// TIA Portal project "HEAT-1-CADIZ-V24" (V20)

(* hardware
DEVICE "S7-1200 station_1"  S7-1200 Station
   slot 0: "Rack_0"  S7-1200 Rack  Rack  V1.0
   slot 1: "PLC_1"  CPU 1214FC DC/DC/RLY  6ES7 214-1HF40-0XB0  V4.6
   slot 2: "DI 16x24VDC_1"  6ES7 221-1BH32-0XB0  V2.0
   slot 3: "DQ 16xRelay_1"  SM 1222 DQ16 x relay  6ES7 222-1HH32-0XB0  V2.0
   slot 4: "F-DI 8/16x24VDC_1"  SM 1226 F-DI8/16 x 24VDC  6ES7 226-6BA32-0XB0  V2.0
   slot 5: "F-DI 8/16x24VDC_2"  SM 1226 F-DI8/16 x 24VDC  6ES7 226-6BA32-0XB0  V2.0
   slot 6: "F-DQ 4x24VDC_1"  SM 1226 F-DQ4 x 24VDC  6ES7 226-6DA32-0XB0  V2.0
DEVICE "GSD device_1"  GSD.Device.PN
   slot 0: "Rack"  Rack  V1.0
   slot 0: "KRC5"  KUKA.PROFINET 6.0  0x300  V6.0
      slot 0: "KUKA.PROFINET 6.0"  KUKA.PROFINET 6.0
      slot 1: "Interface1"  Interface1
         slot 1: "Port001(XF3)"  Port001(XF3)
         slot 2: "Port002(XF4)"  Port002(XF4)
         slot 3: "Port003(XF5)"  Port003(XF5)
         slot 4: "Port004(XF6)"  Port004(XF6)
   slot 1: "64 safe digital in- and outputs (2.4)_1"  64 safe digital in- and outputs (2.4)  KUKADevF64_2.4
      slot 0: "64 safe digital in- and outputs (2.4)"  64 safe digital in- and outputs (2.4)
   slot 2: "1024 digital in- and outputs_1"  1024 digital in- and outputs  KUKA Device IO1024
      slot 0: "1024 digital in- and outputs"  1024 digital in- and outputs
DEVICE "HMI_1"  KTP1200 Basic PN
   slot 0: "HMI_1"  KTP1200 Basic PN  6AV2 123-2MB03-0AX0  17.0.0.0
   slot 1: "HMI_RT_1"  KTP1200 Basic PN  6AV2 123-2MB03-0AX0  17.0.0.0
   slot 5: "HMI_1.IE_CP_1"  PROFINET Interface  17.0.0.0
      slot 1: "PROFINET Interface_1"  PROFINET Interface
         slot 1: "Port_1"  Port
DEVICE "ET 200SP station_2"  ET 200SP-Station
   slot 0: "Rack_0"  Rack  6ES5 710-8MAx1
   slot 0: "islaparking"  IM 155-6 PN ST  6ES7 155-6AU01-0BN0  V4.2
   slot 1: "DI 16x24VDC ST_1"  DI 16x24VDC ST  6ES7 131-6BH01-0BA0  V0.0
      slot 1: "DI 16x24VDC ST_1"  DI 16x24VDC ST
   slot 2: "DI 8x24VDC ST_1"  DI 8x24VDC ST  6ES7 131-6BF01-0BA0  V0.0
      slot 1: "DI 8x24VDC ST_1"  DI 8x24VDC ST
   slot 3: "DQ 16x24VDC/0.5A ST_1"  DQ 16x24VDC/0.5A ST  6ES7 132-6BH01-0BA0  V0.0
      slot 1: "DQ 16x24VDC/0.5A ST_1"  DQ 16x24VDC/0.5A ST
   slot 4: "DQ 8x24VDC/0.5A ST_1"  DQ 8x24VDC/0.5A ST  6ES7 132-6BF01-0BA0  V0.0
      slot 1: "DQ 8x24VDC/0.5A ST_1"  DQ 8x24VDC/0.5A ST
   slot 5: "Server module_1"  Server module  6ES7 193-6PA00-0AA0  V1.1
      slot 1: "Server module_1"  Server module
   slot 127: "BA 2xRJ45"  BA 2xRJ45  6ES7 193-6AR00-0AA0  V0.0
      slot 1: "Port_1"  X1 P1R  6ES7 193-6AR00-0AA0  V0.0
      slot 2: "Port_2"  X1 P2R  6ES7 193-6AR00-0AA0  V0.0
DEVICE "ET 200SP station_1"  ET 200SP-Station
   slot 0: "Rack_0"  Rack  6ES5 710-8MAx1
   slot 0: "islarobot"  IM 155-6 PN ST  6ES7 155-6AU01-0BN0  V4.2
   slot 1: "DI 16x24VDC ST_1"  DI 16x24VDC ST  6ES7 131-6BH01-0BA0  V0.0
      slot 1: "DI 16x24VDC ST_1"  DI 16x24VDC ST
   slot 2: "DI 8x24VDC ST_1"  DI 8x24VDC ST  6ES7 131-6BF01-0BA0  V0.0
      slot 1: "DI 8x24VDC ST_1"  DI 8x24VDC ST
   slot 3: "DQ 16x24VDC/0.5A ST_1"  DQ 16x24VDC/0.5A ST  6ES7 132-6BH01-0BA0  V0.0
      slot 1: "DQ 16x24VDC/0.5A ST_1"  DQ 16x24VDC/0.5A ST
   slot 4: "DQ 8x24VDC/0.5A ST_1"  DQ 8x24VDC/0.5A ST  6ES7 132-6BF01-0BA0  V0.0
      slot 1: "DQ 8x24VDC/0.5A ST_1"  DQ 8x24VDC/0.5A ST
   slot 5: "Server module_1"  Server module  6ES7 193-6PA00-0AA0  V1.1
      slot 1: "Server module_1"  Server module
   slot 127: "BA 2xRJ45"  BA 2xRJ45  6ES7 193-6AR00-0AA0  V0.0
      slot 1: "Port_1"  X1 P1R  6ES7 193-6AR00-0AA0  V0.0
      slot 2: "Port_2"  X1 P2R  6ES7 193-6AR00-0AA0  V0.0
DEVICE "GSD device_2"  GSD.Device.PN
   slot 0: "Rack"  Rack  V1.0
   slot 0: "CPX"  CPX Rev 50  TN 197330
      slot 0: "CPX Rev 50"  CPX Rev 50
      slot 1: "PN-IO Interface"  PN-IO Interface
         slot 1: "Port 1"  Port 1
         slot 2: "Port 2"  Port 2
   slot 1: "FB43 PNIO Module_1"  FB43 PNIO Module  TN 8110369, CPX-FB43
      slot 0: "FB43 PNIO Module"  FB43 PNIO Module
   slot 2: "MPAL DIL 4 [32DO]_1"  MPAL DIL 4 [32DO]
      slot 0: "MPAL DIL 4 [32DO]"  MPAL DIL 4 [32DO]
DEVICE "ET 200SP station_3"  ET 200SP-Station
   slot 0: "Rack_0"  Rack  6ES5 710-8MAx1
   slot 0: "sistemadeagua"  IM 155-6 PN ST  6ES7 155-6AU01-0BN0  V4.2
   slot 1: "DI 8x24VDC ST_1"  DI 8x24VDC ST  6ES7 131-6BF01-0BA0  V0.0
      slot 1: "DI 8x24VDC ST_1"  DI 8x24VDC ST
   slot 2: "DQ 8x24VDC/0.5A ST_1"  DQ 8x24VDC/0.5A ST  6ES7 132-6BF01-0BA0  V0.0
      slot 1: "DQ 8x24VDC/0.5A ST_1"  DQ 8x24VDC/0.5A ST
   slot 3: "AI 4xU/I 2-wire ST_1"  AI 4xU/I 2-wire ST  6ES7 134-6HD01-0BA1  V2.0
      slot 1: "AI 4xU/I 2-wire ST_1"  AI 4xU/I 2-wire ST
   slot 4: "Server module_1"  Server module  6ES7 193-6PA00-0AA0  V1.1
      slot 1: "Server module_1"  Server module
   slot 127: "BA 2xRJ45"  BA 2xRJ45  6ES7 193-6AR00-0AA0  V0.0
      slot 1: "Port_1"  X1 P1R  6ES7 193-6AR00-0AA0  V0.0
      slot 2: "Port_2"  X1 P2R  6ES7 193-6AR00-0AA0  V0.0
DEVICE "GSD device_3"  GSD.Device.PN
   slot 0: "Rack"  Rack  V1.0
   slot 0: "CPX_1"  CPX Rev 50  TN 197330
      slot 0: "CPX Rev 50"  CPX Rev 50
      slot 1: "PN-IO Interface"  PN-IO Interface
         slot 1: "Port 1"  Port 1
         slot 2: "Port 2"  Port 2
   slot 1: "FB43 PNIO Module_1"  FB43 PNIO Module  TN 8110369, CPX-FB43
      slot 0: "FB43 PNIO Module"  FB43 PNIO Module
   slot 2: "16DI [16DI]_1"  16DI [16DI]
      slot 0: "16DI [16DI]"  16DI [16DI]
   slot 3: "16DI [16DI]_2"  16DI [16DI]
      slot 0: "16DI [16DI]"  16DI [16DI]
   slot 4: "MPAL DIL 4 [32DO]_1"  MPAL DIL 4 [32DO]
      slot 0: "MPAL DIL 4 [32DO]"  MPAL DIL 4 [32DO]
*)

// ===== PLC "PLC_1"  CPU 1214FC DC/DC/RLY =====

VAR_GLOBAL   // PLC tag table "Default tag table"
   "RES1 (reservado)" AT %Q500.0 : Bool;
   "eStopButtonCabinet" AT %I40.0 : Bool;   // Emergency-Stop cabinet — 1oo2 result
   "eStopButtonTank" AT %I40.1 : Bool;   // Emergency-Stop tank — 1oo2 result
   "eStopButtonTankPartnerCh" AT %I41.1 : Bool;   // partner channel 1oo2 — do not use
   "eStopButtonWaterSystem" AT %I40.2 : Bool;   // Emergency-Stop water system — 1oo2 result
   "eStopButtonWaterSystemPartnerCh" AT %I41.2 : Bool;   // partner channel 1oo2 — do not use
   "eStopButtonHmiPanel" AT %I40.3 : Bool;   // Emergency-Stop HMI panel — 1oo2 result
   "eStopButtonHmiPanelPartnerCh" AT %I41.3 : Bool;   // partner channel 1oo2 — do not use
   "eStopButtonLightCurtain1" AT %I40.4 : Bool;   // Emergency-Stop light curtain 1 — 1oo2 resul
   "eStopButtonLightCurtain1PartnerCh" AT %I41.4 : Bool;   // partner channel 1oo2 — do not use
   "eStopButtonDoor" AT %I40.5 : Bool;   // Emergency-Stop Door — 1oo2 result
   "eStopButtonDoorPartnerCh" AT %I41.5 : Bool;   // partner channel 1oo2 — do not use
   "lightCurtain1Ossd1" AT %I50.0 : Bool;   // Z2 – LC 1 OSSD 1 (receiver)
   "lightCurtain1Ossd2" AT %I51.0 : Bool;   // Z2 – LC 1 OSSD 2 (receiver)
   "lightCurtain3Ossd1" AT %I50.1 : Bool;   // Z2 – LC 3 OSSD 1 (receiver)
   "lightCurtain3Ossd2" AT %I51.1 : Bool;   // Z2 – LC 3 OSSD 2 (receiver)
   "lightCurtain6Ossd1" AT %I50.2 : Bool;   // Z2 – LC 6 OSSD 1 (receiver)
   "lightCurtain6Ossd2" AT %I51.2 : Bool;   // Z2 – LC 6 OSSD 2 (receiver)
   "enableAccessReqSelector" AT %I50.3 : Bool;   // Rotary selector – enabless request access
   "DoorClosedCh1" AT %I50.6 : Bool;   // Safety door closed interlock – contact 1
   "resetDoorButton" AT %I50.7 : Bool;   // Reset push‑button
   "SAF_DOOR_CLSD_CH2" AT %I51.6 : Bool;   // Safety door closed interlock – contact 2
   "SAF_DOOR_UNLOCK_CH1" AT %Q60.0 : Bool;   // Unlock safety door – redundant output 1
   "SAF_GATE_UNLOCK_CH2" AT %Q60.2 : Bool;   // Unlock safety door – redundant output 2
   "IND_RESET_LAMP" AT %Q10.0 : Bool;   // Reset indicator lamp
   "IND_STATUS_LAMP" AT %Q10.1 : Bool;   // System-status pilot light
   "CMD_PRESS_EXH_VALVE" AT %Q11.0 : Bool;   // Pressure/exhaust solenoid-valve command
   "STS_RECIRC_PUMP" AT %I20.0 : Bool;   // Recirculation-pump feedback
   "STS_TRANSFER_PUMP" AT %I20.1 : Bool;   // Transfer-pump feedback
   "ALM_UV_FILTER" AT %I20.2 : Bool;   // UV-filter fault alarm
   "ALM_PIT_LVL_LOW" AT %I20.3 : Bool;   // Sump low-level alarm
   "ALM_TANK_LVL_LOW" AT %I20.4 : Bool;   // Tank low-level alarm
   "STS_TANK_FILLING" AT %I20.5 : Bool;   // Tank filling status
   "STS_TANK_DRAINING" AT %I20.6 : Bool;   // Tank draining status
   "MODE_WATER_AUTO" AT %Q30.3 : Bool;   // CONMUTADOR AUTO
   "IND_BEACON2_GREEN" AT %Q30.4 : Bool;   // Beacon 2 – green
   "IND_BEACON2_RED" AT %Q30.5 : Bool;   // Beacon 2 – red
   "robotPresenceSignalZone1" AT %I500.0 : Bool;
   "robotPresenceSignalZone2" AT %I500.1 : Bool;
   "robotPresenceSignalZone3" AT %I500.2 : Bool;
   "eStopButtonCabinetPartnerCh" AT %I41.0 : Bool;   // partner channel 1oo2 — do not use
   "lightCurtain2Ossd1" AT %I300.0 : Bool;
   "lightCurtain2Ossd2" AT %I300.4 : Bool;
   "eStopButtonIslandRightPartner" AT %I300.5 : Bool;
   "lightCurtain4Ossd1" AT %I350.0 : Bool;
   "eStopButtonIslandLeft" AT %I350.1 : Bool;
   "lightCurtain5Ossd1" AT %I350.2 : Bool;
   "eStopButtonIslandLefttPartner" AT %I350.3 : Bool;   // partner channel 1oo2 — do not use
   "lightCurtain4Ossd2" AT %I350.4 : Bool;
   "lightCurtain5Ossd2" AT %I350.6 : Bool;
   "accessReqButtonZone2" AT %I51.4 : Bool;   // Illuminated push-button – access request for zone 2
   "accessReqButtonZone3" AT %I51.5 : Bool;   // Illuminated push-button – access request for zone 3
   "accessReqButtonZone1" AT %I51.3 : Bool;   // Illuminated push-button – access request for zone 1
   "eStopButtonIslandRight" AT %I300.1 : Bool;
   "NHE – E‑Stop externo  NO pulsado" AT %Q500.1 : Bool;
   "BS – Puerta cerrada" AT %Q500.2 : Bool;
   "QBS – Ack puerta" AT %Q500.3 : Bool;
   "SHS1 – Stop 1" AT %Q500.4 : Bool;
   "SHS2 – Stop 2" AT %Q500.5 : Bool;
   "RES6" AT %Q500.6 : Bool;
   "RES7" AT %Q500.7 : Bool;
   "US2 – 24 V US2" AT %Q501.0 : Bool;
   "SBH – Safe Op Stop" AT %Q501.1 : Bool;
   "RES11" AT %Q501.2 : Bool;
   "RES12" AT %Q501.3 : Bool;
   "RES13" AT %Q501.4 : Bool;
   "RES14" AT %Q501.5 : Bool;
   "RES15" AT %Q501.6 : Bool;
   "SPA – Power‑down Ack" AT %Q501.7 : Bool;
   "resetHmiButton" AT %I51.7 : Bool;
   "Tag_1" AT %M200.0 : Bool;
   "Tag_2" AT %M201.0 : Bool;
   "Tag_3" AT %M500.1 : Bool;
   "Tag_4" AT %M755.5 : Bool;
   "V5" AT %Q0.4 : Bool;   // Biestable_B_RETROCESO
   "ABRIR_TAPA_PEPA" AT %Q170.2 : Bool;
   "CERRAR_TAPA_PEPA" AT %Q170.3 : Bool;
   "ABRIR_TAPA_INMERSION" AT %Q170.4 : Bool;
   "CERRAR_TAPA_INMERSION" AT %Q170.5 : Bool;
   "ABRIR_TAPA_MARCADOR" AT %Q170.6 : Bool;
   "CERRAR_TAPA_MARCADOR" AT %Q170.7 : Bool;
   "ABRIR_TAPA_PERFILOMETRO" AT %Q171.0 : Bool;
   "CERRAR_TAPA_PERFILOMETRO" AT %Q171.1 : Bool;
   "V6" AT %Q0.5 : Bool;   // Biestable_A_AVANCE
   "V7" AT %Q0.6 : Bool;
   "V8" AT %Q0.7 : Bool;
   "moveCode_00" AT %Q616.0 : Bool;
   "goTrigger" AT %Q622.0 : Bool;
   "baseReqId_00" AT %Q620.0 : Bool;
   "baseReqId_01" AT %Q620.1 : Bool;
   "baseReqId_02" AT %Q620.2 : Bool;
   "baseReqId_03" AT %Q620.3 : Bool;
   "baseReqId_04" AT %Q620.4 : Bool;
   "baseReqId_05" AT %Q620.5 : Bool;
   "baseReqId_06" AT %Q620.6 : Bool;
   "baseReqId_07" AT %Q620.7 : Bool;
   "baseReqId_08" AT %Q621.0 : Bool;
   "baseReqId_09" AT %Q621.1 : Bool;
   "baseReqId_10" AT %Q621.2 : Bool;
   "baseReqId_11" AT %Q621.3 : Bool;
   "baseReqId_12" AT %Q621.4 : Bool;
   "baseReqId_13" AT %Q621.5 : Bool;
   "baseReqId_14" AT %Q621.6 : Bool;
   "baseReqId_15" AT %Q621.7 : Bool;
   "moveCode_01" AT %Q616.1 : Bool;
   "moveCode_02" AT %Q616.2 : Bool;
   "moveCode_03" AT %Q616.3 : Bool;
   "moveCode_04" AT %Q616.4 : Bool;
   "moveCode_05" AT %Q616.5 : Bool;
   "moveCode_06" AT %Q616.6 : Bool;
   "moveCode_07" AT %Q616.7 : Bool;
   "moveCode_08" AT %Q617.0 : Bool;
   "moveCode_09" AT %Q617.1 : Bool;
   "moveCode_10" AT %Q617.2 : Bool;
   "moveCode_11" AT %Q617.3 : Bool;
   "moveCode_12" AT %Q617.4 : Bool;
   "moveCode_13" AT %Q617.5 : Bool;
   "moveCode_14" AT %Q617.6 : Bool;
   "moveCode_15" AT %Q617.7 : Bool;
   "toolNo_00" AT %I625.0 : Bool;
   "toolNo_01" AT %I625.1 : Bool;
   "toolNo_02" AT %I625.2 : Bool;
   "toolNo_03" AT %I625.3 : Bool;
   "toolNo_04" AT %I625.4 : Bool;
   "toolNo_05" AT %I625.5 : Bool;
   "toolNo_06" AT %I625.6 : Bool;
   "toolNo_07" AT %I625.7 : Bool;
   "baseNo_00" AT %I626.0 : Bool;
   "baseNo_01" AT %I626.1 : Bool;
   "baseNo_02" AT %I626.2 : Bool;
   "baseNo_03" AT %I626.3 : Bool;
   "baseNo_04" AT %I626.4 : Bool;
   "baseNo_05" AT %I626.5 : Bool;
   "baseNo_06" AT %I626.6 : Bool;
   "baseNo_07" AT %I626.7 : Bool;
   "toolNoByte" AT %IB625 : Byte;
   "baseNoByte" AT %IB626 : Byte;
   "programReqId_00" AT %Q623.0 : Bool;
   "programReqId_01" AT %Q623.1 : Bool;
   "programReqId_02" AT %Q623.2 : Bool;
   "programReqId_03" AT %Q623.3 : Bool;
   "programReqId_04" AT %Q623.4 : Bool;
   "programReqId_05" AT %Q623.5 : Bool;
   "programReqId_06" AT %Q623.6 : Bool;
   "programReqId_07" AT %Q623.7 : Bool;
   "programReqId_08" AT %Q624.0 : Bool;
   "programReqId_09" AT %Q624.1 : Bool;
   "programReqId_10" AT %Q624.2 : Bool;
   "programReqId_11" AT %Q624.3 : Bool;
   "programReqId_12" AT %Q624.4 : Bool;
   "programReqId_13" AT %Q624.5 : Bool;
   "programReqId_14" AT %Q624.6 : Bool;
   "programReqId_15" AT %Q624.7 : Bool;
   "programReqId" AT %QW623 : Word;
   "PRUEBA_4" AT %Q4.4 : Bool;
   "PRUEBA_5" AT %Q4.5 : Bool;
   "PRUEBA_JOAQUIN" AT %Q4.0 : Bool;
   "PRUEBA_6" AT %Q4.6 : Bool;
   "PRUEBA_7" AT %Q4.7 : Bool;
   "cancelGo" AT %Q625.0 : Bool;
   "pauseGo" AT %Q625.1 : Bool;
   "resumeGo" AT %Q625.2 : Bool;
   "ACTIVAR_AGUA" AT %Q220.1 : Bool;   // VALVULA EMBARCADA ISLA ROBOT
   "AGUA_JOAQUIN" AT %Q4.3 : Bool;   // SISTEMA DE AGUA - JOAQUIN
   "PGNO_BIT_00" AT %Q626.0 : Bool;   // $IN[209] en KUKA
   "PGNO_BIT_01" AT %Q626.1 : Bool;   // $IN[210] en KUKA
   "PGNO_BIT_02" AT %Q626.2 : Bool;   // $IN[211] en KUKA
   "PGNO_BIT_03" AT %Q626.3 : Bool;
   "PGNO_BIT_04" AT %Q626.4 : Bool;
   "PGNO_BIT_05" AT %Q626.5 : Bool;
   "PGNO_BIT_06" AT %Q626.6 : Bool;
   "PGNO_BIT_07" AT %Q626.7 : Bool;
   "PGNO_PARITY" AT %Q627.0 : Bool;   // $IN[217] en KUKA
   "PGNO_VALID" AT %Q627.1 : Bool;   // $IN[218] en KUKA
   "$EXT_START" AT %Q627.2 : Bool;   // $IN[219] en KUKA
   "$MOVE_ENABLE" AT %Q627.3 : Bool;   // $IN[220] en KUKA
   "$CONF_MESS" AT %Q627.4 : Bool;   // $IN[221] en KUKA
   "$DRIVES_OFF" AT %Q627.5 : Bool;   // $IN[222] en KUKA
   "$DRIVES_ON" AT %Q627.6 : Bool;   // $IN[223] en KUKA
   "$I_O_ACT" AT %Q627.7 : Bool;   // $IN[224] en KUKA
   "PGNO_REQ" AT %I624.7 : Bool;   // OUT[200] EN KUKA
   "startAutoExt" AT %M777.0 : Bool;
   "Tag_6" AT %Q220.0 : Bool;
   "Tag_7" AT %Q4.1 : Bool;
   "Tag_8" AT %Q4.2 : Bool;
   "Tag_9" AT %I0.4 : Bool;
   "Tag_10" AT %I0.0 : Bool;
   "Tag_11" AT %I0.1 : Bool;
   "Tag_12" AT %I0.2 : Bool;
   "Tag_13" AT %I0.3 : Bool;
   "Tag_14" AT %I210.1 : Bool;
   "Tag_15" AT %I210.2 : Bool;
   "Tag_16" AT %I210.0 : Bool;
   "Tag_17" AT %I210.3 : Bool;
   "Tag_18" AT %I210.4 : Bool;
   "AchimHmiEnable" AT %M202.0 : Bool;
   "toolIdProxy1" AT %I201.3 : Bool;
   "toolIdProxy2" AT %I201.2 : Bool;
   "toolIdProxy3" AT %I201.1 : Bool;
   "toolIdProxy4" AT %I201.0 : Bool;
   "dockValveV2UnlockOnPole" AT %Q171.6 : Bool;
   "$PRO_ACT" AT %I627.2 : Bool;   // OUT[219] EN KUKA
   "$STOPMESS" AT %I627.1 : Bool;   // OUT[218] EN KUKA
   "$PERI_RDY" AT %I627.0 : Bool;   // OUT[217] EN KUKA
   "robotInLoopKukaControl" AT %Q628.0 : Bool;
   "robotInLoopSupervisor" AT %Q628.1 : Bool;
   "xInicial_00" AT %Q632.0 : Bool;
   "xInicial_01" AT %Q632.1 : Bool;
   "xInicial_02" AT %Q632.2 : Bool;
   "xInicial_03" AT %Q632.3 : Bool;
   "xInicial_04" AT %Q632.4 : Bool;
   "xInicial_05" AT %Q632.5 : Bool;
   "xInicial_06" AT %Q632.6 : Bool;
   "xInicial_07" AT %Q632.7 : Bool;
   "xInicial_08" AT %Q633.0 : Bool;
   "xInicial_09" AT %Q633.1 : Bool;
   "xInicial_10" AT %Q633.2 : Bool;
   "xInicial_11" AT %Q633.3 : Bool;
   "xInicial_12" AT %Q633.4 : Bool;
   "xInicial_13" AT %Q633.5 : Bool;
   "xInicial_14" AT %Q633.6 : Bool;
   "xInicial_15" AT %Q633.7 : Bool;
   "xInicial_16" AT %Q634.0 : Bool;
   "xInicial_17" AT %Q634.1 : Bool;
   "xInicial_18" AT %Q634.2 : Bool;
   "xInicial_19" AT %Q634.3 : Bool;
   "xInicial_20" AT %Q634.4 : Bool;
   "xInicial_21" AT %Q634.5 : Bool;
   "xInicial_22" AT %Q634.6 : Bool;
   "xInicial_23" AT %Q634.7 : Bool;
   "xInicial_24" AT %Q635.0 : Bool;
   "xInicial_25" AT %Q635.1 : Bool;
   "xInicial_26" AT %Q635.2 : Bool;
   "xInicial_27" AT %Q635.3 : Bool;
   "xInicial_28" AT %Q635.4 : Bool;
   "xInicial_29" AT %Q635.5 : Bool;
   "xInicial_30" AT %Q635.6 : Bool;
   "xInicial_31" AT %Q635.7 : Bool;
   "yInicial_00" AT %Q636.0 : Bool;
   "yInicial_01" AT %Q636.1 : Bool;
   "yInicial_02" AT %Q636.2 : Bool;
   "yInicial_03" AT %Q636.3 : Bool;
   "yInicial_04" AT %Q636.4 : Bool;
   "yInicial_05" AT %Q636.5 : Bool;
   "yInicial_06" AT %Q636.6 : Bool;
   "yInicial_07" AT %Q636.7 : Bool;
   "yInicial_08" AT %Q637.0 : Bool;
   "yInicial_09" AT %Q637.1 : Bool;
   "yInicial_10" AT %Q637.2 : Bool;
   "yInicial_11" AT %Q637.3 : Bool;
   "yInicial_12" AT %Q637.4 : Bool;
   "yInicial_13" AT %Q637.5 : Bool;
   "yInicial_14" AT %Q637.6 : Bool;
   "yInicial_15" AT %Q637.7 : Bool;
   "yInicial_16" AT %Q638.0 : Bool;
   "yInicial_17" AT %Q638.1 : Bool;
   "yInicial_18" AT %Q638.2 : Bool;
   "yInicial_19" AT %Q638.3 : Bool;
   "yInicial_20" AT %Q638.4 : Bool;
   "yInicial_21" AT %Q638.5 : Bool;
   "yInicial_22" AT %Q638.6 : Bool;
   "yInicial_23" AT %Q638.7 : Bool;
   "yInicial_24" AT %Q639.0 : Bool;
   "yInicial_25" AT %Q639.1 : Bool;
   "yInicial_26" AT %Q639.2 : Bool;
   "yInicial_27" AT %Q639.3 : Bool;
   "yInicial_28" AT %Q639.4 : Bool;
   "yInicial_29" AT %Q639.5 : Bool;
   "yInicial_30" AT %Q639.6 : Bool;
   "yInicial_31" AT %Q639.7 : Bool;
   "zInicial_00" AT %Q640.0 : Bool;
   "zInicial_01" AT %Q640.1 : Bool;
   "zInicial_02" AT %Q640.2 : Bool;
   "zInicial_03" AT %Q640.3 : Bool;
   "zInicial_04" AT %Q640.4 : Bool;
   "zInicial_05" AT %Q640.5 : Bool;
   "zInicial_06" AT %Q640.6 : Bool;
   "zInicial_07" AT %Q640.7 : Bool;
   "zInicial_08" AT %Q641.0 : Bool;
   "zInicial_09" AT %Q641.1 : Bool;
   "zInicial_10" AT %Q641.2 : Bool;
   "zInicial_11" AT %Q641.3 : Bool;
   "zInicial_12" AT %Q641.4 : Bool;
   "zInicial_13" AT %Q641.5 : Bool;
   "zInicial_14" AT %Q641.6 : Bool;
   "zInicial_15" AT %Q641.7 : Bool;
   "zInicial_16" AT %Q642.0 : Bool;
   "zInicial_17" AT %Q642.1 : Bool;
   "zInicial_18" AT %Q642.2 : Bool;
   "zInicial_19" AT %Q642.3 : Bool;
   "zInicial_20" AT %Q642.4 : Bool;
   "zInicial_21" AT %Q642.5 : Bool;
   "zInicial_22" AT %Q642.6 : Bool;
   "zInicial_23" AT %Q642.7 : Bool;
   "zInicial_24" AT %Q643.0 : Bool;
   "zInicial_25" AT %Q643.1 : Bool;
   "zInicial_26" AT %Q643.2 : Bool;
   "zInicial_27" AT %Q643.3 : Bool;
   "zInicial_28" AT %Q643.4 : Bool;
   "zInicial_29" AT %Q643.5 : Bool;
   "zInicial_30" AT %Q643.6 : Bool;
   "zInicial_31" AT %Q643.7 : Bool;
   "e1Inicial_00" AT %Q644.0 : Bool;
   "e1Inicial_01" AT %Q644.1 : Bool;
   "e1Inicial_02" AT %Q644.2 : Bool;
   "e1Inicial_03" AT %Q644.3 : Bool;
   "e1Inicial_04" AT %Q644.4 : Bool;
   "e1Inicial_05" AT %Q644.5 : Bool;
   "e1Inicial_06" AT %Q644.6 : Bool;
   "e1Inicial_07" AT %Q644.7 : Bool;
   "e1Inicial_08" AT %Q645.0 : Bool;
   "e1Inicial_09" AT %Q645.1 : Bool;
   "e1Inicial_10" AT %Q645.2 : Bool;
   "e1Inicial_11" AT %Q645.3 : Bool;
   "e1Inicial_12" AT %Q645.4 : Bool;
   "e1Inicial_13" AT %Q645.5 : Bool;
   "e1Inicial_14" AT %Q645.6 : Bool;
   "e1Inicial_15" AT %Q645.7 : Bool;
   "e1Inicial_16" AT %Q646.0 : Bool;
   "e1Inicial_17" AT %Q646.1 : Bool;
   "e1Inicial_18" AT %Q646.2 : Bool;
   "e1Inicial_19" AT %Q646.3 : Bool;
   "e1Inicial_20" AT %Q646.4 : Bool;
   "e1Inicial_21" AT %Q646.5 : Bool;
   "e1Inicial_22" AT %Q646.6 : Bool;
   "e1Inicial_23" AT %Q646.7 : Bool;
   "e1Inicial_24" AT %Q647.0 : Bool;
   "e1Inicial_25" AT %Q647.1 : Bool;
   "e1Inicial_26" AT %Q647.2 : Bool;
   "e1Inicial_27" AT %Q647.3 : Bool;
   "e1Inicial_28" AT %Q647.4 : Bool;
   "e1Inicial_29" AT %Q647.5 : Bool;
   "e1Inicial_30" AT %Q647.6 : Bool;
   "e1Inicial_31" AT %Q647.7 : Bool;
   "xFinal_00" AT %Q648.0 : Bool;
   "xFinal_01" AT %Q648.1 : Bool;
   "xFinal_02" AT %Q648.2 : Bool;
   "xFinal_03" AT %Q648.3 : Bool;
   "xFinal_04" AT %Q648.4 : Bool;
   "xFinal_05" AT %Q648.5 : Bool;
   "xFinal_06" AT %Q648.6 : Bool;
   "xFinal_07" AT %Q648.7 : Bool;
   "xFinal_08" AT %Q649.0 : Bool;
   "xFinal_09" AT %Q649.1 : Bool;
   "xFinal_10" AT %Q649.2 : Bool;
   "xFinal_11" AT %Q649.3 : Bool;
   "xFinal_12" AT %Q649.4 : Bool;
   "xFinal_13" AT %Q649.5 : Bool;
   "xFinal_14" AT %Q649.6 : Bool;
   "xFinal_15" AT %Q649.7 : Bool;
   "xFinal_16" AT %Q650.0 : Bool;
   "xFinal_17" AT %Q650.1 : Bool;
   "xFinal_18" AT %Q650.2 : Bool;
   "xFinal_19" AT %Q650.3 : Bool;
   "xFinal_20" AT %Q650.4 : Bool;
   "xFinal_21" AT %Q650.5 : Bool;
   "xFinal_22" AT %Q650.6 : Bool;
   "xFinal_23" AT %Q650.7 : Bool;
   "xFinal_24" AT %Q651.0 : Bool;
   "xFinal_25" AT %Q651.1 : Bool;
   "xFinal_26" AT %Q651.2 : Bool;
   "xFinal_27" AT %Q651.3 : Bool;
   "xFinal_28" AT %Q651.4 : Bool;
   "xFinal_29" AT %Q651.5 : Bool;
   "xFinal_30" AT %Q651.6 : Bool;
   "xFinal_31" AT %Q651.7 : Bool;
   "yFinal_00" AT %Q652.0 : Bool;
   "yFinal_01" AT %Q652.1 : Bool;
   "yFinal_02" AT %Q652.2 : Bool;
   "yFinal_03" AT %Q652.3 : Bool;
   "yFinal_04" AT %Q652.4 : Bool;
   "yFinal_05" AT %Q652.5 : Bool;
   "yFinal_06" AT %Q652.6 : Bool;
   "yFinal_07" AT %Q652.7 : Bool;
   "yFinal_08" AT %Q653.0 : Bool;
   "yFinal_09" AT %Q653.1 : Bool;
   "yFinal_10" AT %Q653.2 : Bool;
   "yFinal_11" AT %Q653.3 : Bool;
   "yFinal_12" AT %Q653.4 : Bool;
   "yFinal_13" AT %Q653.5 : Bool;
   "yFinal_14" AT %Q653.6 : Bool;
   "yFinal_15" AT %Q653.7 : Bool;
   "yFinal_16" AT %Q654.0 : Bool;
   "yFinal_17" AT %Q654.1 : Bool;
   "yFinal_18" AT %Q654.2 : Bool;
   "yFinal_19" AT %Q654.3 : Bool;
   "yFinal_20" AT %Q654.4 : Bool;
   "yFinal_21" AT %Q654.5 : Bool;
   "yFinal_22" AT %Q654.6 : Bool;
   "yFinal_23" AT %Q654.7 : Bool;
   "yFinal_24" AT %Q655.0 : Bool;
   "yFinal_25" AT %Q655.1 : Bool;
   "yFinal_26" AT %Q655.2 : Bool;
   "yFinal_27" AT %Q655.3 : Bool;
   "yFinal_28" AT %Q655.4 : Bool;
   "yFinal_29" AT %Q655.5 : Bool;
   "yFinal_30" AT %Q655.6 : Bool;
   "yFinal_31" AT %Q655.7 : Bool;
   "zFinal_00" AT %Q656.0 : Bool;
   "zFinal_01" AT %Q656.1 : Bool;
   "zFinal_02" AT %Q656.2 : Bool;
   "zFinal_03" AT %Q656.3 : Bool;
   "zFinal_04" AT %Q656.4 : Bool;
   "zFinal_05" AT %Q656.5 : Bool;
   "zFinal_06" AT %Q656.6 : Bool;
   "zFinal_07" AT %Q656.7 : Bool;
   "zFinal_08" AT %Q657.0 : Bool;
   "zFinal_09" AT %Q657.1 : Bool;
   "zFinal_10" AT %Q657.2 : Bool;
   "zFinal_11" AT %Q657.3 : Bool;
   "zFinal_12" AT %Q657.4 : Bool;
   "zFinal_13" AT %Q657.5 : Bool;
   "zFinal_14" AT %Q657.6 : Bool;
   "zFinal_15" AT %Q657.7 : Bool;
   "zFinal_16" AT %Q658.0 : Bool;
   "zFinal_17" AT %Q658.1 : Bool;
   "zFinal_18" AT %Q658.2 : Bool;
   "zFinal_19" AT %Q658.3 : Bool;
   "zFinal_20" AT %Q658.4 : Bool;
   "zFinal_21" AT %Q658.5 : Bool;
   "zFinal_22" AT %Q658.6 : Bool;
   "zFinal_23" AT %Q658.7 : Bool;
   "zFinal_24" AT %Q659.0 : Bool;
   "zFinal_25" AT %Q659.1 : Bool;
   "zFinal_26" AT %Q659.2 : Bool;
   "zFinal_27" AT %Q659.3 : Bool;
   "zFinal_28" AT %Q659.4 : Bool;
   "zFinal_29" AT %Q659.5 : Bool;
   "zFinal_30" AT %Q659.6 : Bool;
   "zFinal_31" AT %Q659.7 : Bool;
   "e1Final_00" AT %Q660.0 : Bool;
   "e1Final_01" AT %Q660.1 : Bool;
   "e1Final_02" AT %Q660.2 : Bool;
   "e1Final_03" AT %Q660.3 : Bool;
   "e1Final_04" AT %Q660.4 : Bool;
   "e1Final_05" AT %Q660.5 : Bool;
   "e1Final_06" AT %Q660.6 : Bool;
   "e1Final_07" AT %Q660.7 : Bool;
   "e1Final_08" AT %Q661.0 : Bool;
   "e1Final_09" AT %Q661.1 : Bool;
   "e1Final_10" AT %Q661.2 : Bool;
   "e1Final_11" AT %Q661.3 : Bool;
   "e1Final_12" AT %Q661.4 : Bool;
   "e1Final_13" AT %Q661.5 : Bool;
   "e1Final_14" AT %Q661.6 : Bool;
   "e1Final_15" AT %Q661.7 : Bool;
   "e1Final_16" AT %Q662.0 : Bool;
   "e1Final_17" AT %Q662.1 : Bool;
   "e1Final_18" AT %Q662.2 : Bool;
   "e1Final_19" AT %Q662.3 : Bool;
   "e1Final_20" AT %Q662.4 : Bool;
   "e1Final_21" AT %Q662.5 : Bool;
   "e1Final_22" AT %Q662.6 : Bool;
   "e1Final_23" AT %Q662.7 : Bool;
   "e1Final_24" AT %Q663.0 : Bool;
   "e1Final_25" AT %Q663.1 : Bool;
   "e1Final_26" AT %Q663.2 : Bool;
   "e1Final_27" AT %Q663.3 : Bool;
   "e1Final_28" AT %Q663.4 : Bool;
   "e1Final_29" AT %Q663.5 : Bool;
   "e1Final_30" AT %Q663.6 : Bool;
   "e1Final_31" AT %Q663.7 : Bool;
   "velRequest_00" AT %Q664.0 : Bool;
   "velRequest_01" AT %Q664.1 : Bool;
   "velRequest_02" AT %Q664.2 : Bool;
   "velRequest_03" AT %Q664.3 : Bool;
   "velRequest_04" AT %Q664.4 : Bool;
   "velRequest_05" AT %Q664.5 : Bool;
   "velRequest_06" AT %Q664.6 : Bool;
   "velRequest_07" AT %Q664.7 : Bool;
   "velRequest_08" AT %Q665.0 : Bool;
   "velRequest_09" AT %Q665.1 : Bool;
   "velRequest_10" AT %Q665.2 : Bool;
   "velRequest_11" AT %Q665.3 : Bool;
   "velRequest_12" AT %Q665.4 : Bool;
   "velRequest_13" AT %Q665.5 : Bool;
   "velRequest_14" AT %Q665.6 : Bool;
   "velRequest_15" AT %Q665.7 : Bool;
   "indexRequest_00" AT %Q666.0 : Bool;
   "indexRequest_01" AT %Q666.1 : Bool;
   "indexRequest_02" AT %Q666.2 : Bool;
   "indexRequest_03" AT %Q666.3 : Bool;
   "indexRequest_04" AT %Q666.4 : Bool;
   "indexRequest_05" AT %Q666.5 : Bool;
   "indexRequest_06" AT %Q666.6 : Bool;
   "indexRequest_07" AT %Q666.7 : Bool;
   "indexRequest_08" AT %Q667.0 : Bool;
   "indexRequest_09" AT %Q667.1 : Bool;
   "indexRequest_10" AT %Q667.2 : Bool;
   "indexRequest_11" AT %Q667.3 : Bool;
   "indexRequest_12" AT %Q667.4 : Bool;
   "indexRequest_13" AT %Q667.5 : Bool;
   "indexRequest_14" AT %Q667.6 : Bool;
   "indexRequest_15" AT %Q667.7 : Bool;
   "Tag_5" AT %M1000.1 : Bool;
   "toolInRobot_00" AT %Q668.0 : Bool;
   "toolInRobot_01" AT %Q668.1 : Bool;
   "toolInRobot_02" AT %Q668.2 : Bool;
   "toolInRobot_03" AT %Q668.3 : Bool;
   "toolInRobot_04" AT %Q668.4 : Bool;
   "toolInRobot_05" AT %Q668.5 : Bool;
   "toolInRobot_06" AT %Q668.6 : Bool;
   "toolInRobot_07" AT %Q668.7 : Bool;
   "kukaFeedBackToolInRobot" AT %QW668 : Word;
   "toolInRobot_08" AT %Q669.0 : Bool;
   "toolInRobot_09" AT %Q669.1 : Bool;
   "toolInRobot_10" AT %Q669.2 : Bool;
   "toolInRobot_11" AT %Q669.3 : Bool;
   "toolInRobot_12" AT %Q669.4 : Bool;
   "toolInRobot_13" AT %Q669.5 : Bool;
   "toolInRobot_14" AT %Q669.6 : Bool;
   "toolInRobot_15" AT %Q669.7 : Bool;
   "kukaAtPerspexPos" AT %I698.0 : Bool;
   "kukaAtGainPos" AT %I698.1 : Bool;
   "kukaAtTcgPos" AT %I698.2 : Bool;
   "kukaAtRefStart" AT %I698.3 : Bool;
   "kukaAtInspStart" AT %I698.4 : Bool;
   "kukaRefScanFin" AT %I698.5 : Bool;
   "kukaInspScanFin" AT %I698.6 : Bool;
   "requestVelocityKuka" AT %QW664 : Word;
   "requestIndexKuka" AT %QW666 : Word;
   "$IN_HOME" AT %I627.3 : Bool;   // OUT[220] EN KUKA
   "$EXT" AT %I627.4 : Bool;   // OUT[221] EN KUKA
END_VAR

VAR_GLOBAL   // PLC tag table "Robot Jog"
   "tcpTargetX_01" AT %Q600.1 : Bool;
   "tcpTargetX_02" AT %Q600.2 : Bool;
   "tcpTargetX_03" AT %Q600.3 : Bool;
   "tcpTargetX_04" AT %Q600.4 : Bool;
   "tcpTargetX_05" AT %Q600.5 : Bool;
   "tcpTargetX_08" AT %Q601.0 : Bool;
   "tcpTargetX_16" AT %Q602.0 : Bool;
   "tcpTargetX_17" AT %Q602.1 : Bool;
   "tcpTargetX_06" AT %Q600.6 : Bool;
   "tcpTargetX_07" AT %Q600.7 : Bool;
   "tcpTargetX_09" AT %Q601.1 : Bool;
   "tcpTargetX_10" AT %Q601.2 : Bool;
   "tcpTargetX_11" AT %Q601.3 : Bool;
   "tcpTargetX_12" AT %Q601.4 : Bool;
   "tcpTargetX_13" AT %Q601.5 : Bool;
   "tcpTargetX_14" AT %Q601.6 : Bool;
   "tcpTargetX_15" AT %Q601.7 : Bool;
   "tcpTargetX_18" AT %Q602.2 : Bool;
   "tcpTargetX_19" AT %Q602.3 : Bool;
   "tcpTargetX_20" AT %Q602.4 : Bool;
   "tcpTargetX_21" AT %Q602.5 : Bool;
   "tcpTargetX_22" AT %Q602.6 : Bool;
   "tcpTargetX_23" AT %Q602.7 : Bool;
   "tcpTargetX_24" AT %Q603.0 : Bool;
   "tcpTargetX_25" AT %Q603.1 : Bool;
   "tcpTargetX_26" AT %Q603.2 : Bool;
   "tcpTargetX_27" AT %Q603.3 : Bool;
   "tcpTargetX_28" AT %Q603.4 : Bool;
   "tcpTargetX_29" AT %Q603.5 : Bool;
   "tcpTargetX_30" AT %Q603.6 : Bool;
   "tcpTargetX_31" AT %Q603.7 : Bool;
   "tcpTargetY_00" AT %Q604.0 : Bool;
   "tcpTargetY_01" AT %Q604.1 : Bool;
   "tcpTargetY_02" AT %Q604.2 : Bool;
   "tcpTargetY_03" AT %Q604.3 : Bool;
   "tcpTargetY_04" AT %Q604.4 : Bool;
   "tcpTargetY_05" AT %Q604.5 : Bool;
   "tcpTargetY_06" AT %Q604.6 : Bool;
   "tcpTargetY_07" AT %Q604.7 : Bool;
   "tcpTargetY_08" AT %Q605.0 : Bool;
   "tcpTargetY_09" AT %Q605.1 : Bool;
   "tcpTargetY_10" AT %Q605.2 : Bool;
   "tcpTargetY_11" AT %Q605.3 : Bool;
   "tcpTargetY_12" AT %Q605.4 : Bool;
   "tcpTargetY_13" AT %Q605.5 : Bool;
   "tcpTargetY_14" AT %Q605.6 : Bool;
   "tcpTargetY_15" AT %Q605.7 : Bool;
   "tcpTargetY_16" AT %Q606.0 : Bool;   // $IN[49]
   "tcpTargetY_17" AT %Q606.1 : Bool;   // $IN[50]
   "tcpTargetY_18" AT %Q606.2 : Bool;   // $IN[51]
   "tcpTargetY_19" AT %Q606.3 : Bool;   // true
   "tcpTargetY_20" AT %Q606.4 : Bool;
   "tcpTargetY_21" AT %Q606.5 : Bool;   // true
   "tcpTargetY_22" AT %Q606.6 : Bool;   // true
   "tcpTargetY_23" AT %Q606.7 : Bool;   // true
   "tcpTargetY_24" AT %Q607.0 : Bool;   // true
   "tcpTargetY_25" AT %Q607.1 : Bool;   // true
   "tcpTargetY_26" AT %Q607.2 : Bool;   // true
   "tcpTargetY_27" AT %Q607.3 : Bool;
   "tcpTargetY_28" AT %Q607.4 : Bool;
   "tcpTargetY_29" AT %Q607.5 : Bool;
   "tcpTargetY_30" AT %Q607.6 : Bool;
   "tcpTargetY_31" AT %Q607.7 : Bool;
   "tcpTargetZ_00" AT %Q608.0 : Bool;
   "tcpTargetZ_01" AT %Q608.1 : Bool;
   "tcpTargetZ_02" AT %Q608.2 : Bool;
   "tcpTargetZ_03" AT %Q608.3 : Bool;
   "tcpTargetZ_04" AT %Q608.4 : Bool;
   "tcpTargetZ_05" AT %Q608.5 : Bool;
   "tcpTargetZ_06" AT %Q608.6 : Bool;
   "tcpTargetZ_07" AT %Q608.7 : Bool;
   "tcpTargetZ_08" AT %Q609.0 : Bool;
   "tcpTargetZ_09" AT %Q609.1 : Bool;
   "tcpTargetZ_10" AT %Q609.2 : Bool;
   "tcpTargetZ_11" AT %Q609.3 : Bool;
   "tcpTargetZ_12" AT %Q609.4 : Bool;
   "tcpTargetZ_13" AT %Q609.5 : Bool;
   "tcpTargetZ_14" AT %Q609.6 : Bool;
   "tcpTargetZ_15" AT %Q609.7 : Bool;
   "tcpTargetZ_16" AT %Q610.0 : Bool;
   "tcpTargetZ_17" AT %Q610.1 : Bool;
   "tcpTargetZ_18" AT %Q610.2 : Bool;
   "tcpTargetZ_19" AT %Q610.3 : Bool;
   "tcpTargetZ_20" AT %Q610.4 : Bool;
   "tcpTargetZ_21" AT %Q610.5 : Bool;
   "tcpTargetZ_22" AT %Q610.6 : Bool;
   "tcpTargetZ_23" AT %Q610.7 : Bool;
   "tcpTargetZ_24" AT %Q611.0 : Bool;
   "tcpTargetZ_25" AT %Q611.1 : Bool;
   "tcpTargetZ_26" AT %Q611.2 : Bool;
   "tcpTargetZ_27" AT %Q611.3 : Bool;
   "tcpTargetZ_28" AT %Q611.4 : Bool;
   "tcpTargetZ_29" AT %Q611.5 : Bool;
   "tcpTargetZ_30" AT %Q611.6 : Bool;
   "tcpTargetZ_31" AT %Q611.7 : Bool;
   "e1Target_00" AT %Q612.0 : Bool;
   "e1Target_01" AT %Q612.1 : Bool;
   "e1Target_02" AT %Q612.2 : Bool;
   "e1Target_03" AT %Q612.3 : Bool;
   "e1Target_04" AT %Q612.4 : Bool;
   "e1Target_05" AT %Q612.5 : Bool;
   "e1Target_06" AT %Q612.6 : Bool;
   "e1Target_07" AT %Q612.7 : Bool;
   "e1Target_08" AT %Q613.0 : Bool;
   "e1Target_09" AT %Q613.1 : Bool;
   "e1Target_10" AT %Q613.2 : Bool;
   "e1Target_11" AT %Q613.3 : Bool;
   "e1Target_12" AT %Q613.4 : Bool;
   "e1Target_13" AT %Q613.5 : Bool;
   "e1Target_14" AT %Q613.6 : Bool;
   "e1Target_15" AT %Q613.7 : Bool;
   "e1Target_16" AT %Q614.0 : Bool;
   "e1Target_17" AT %Q614.1 : Bool;
   "e1Target_18" AT %Q614.2 : Bool;
   "e1Target_19" AT %Q614.3 : Bool;
   "e1Target_20" AT %Q614.4 : Bool;
   "e1Target_21" AT %Q614.5 : Bool;
   "e1Target_22" AT %Q614.6 : Bool;
   "e1Target_23" AT %Q614.7 : Bool;
   "e1Target_24" AT %Q615.0 : Bool;
   "e1Target_25" AT %Q615.1 : Bool;
   "e1Target_26" AT %Q615.2 : Bool;
   "e1Target_27" AT %Q615.3 : Bool;
   "e1Target_28" AT %Q615.4 : Bool;
   "e1Target_29" AT %Q615.5 : Bool;
   "e1Target_30" AT %Q615.6 : Bool;
   "e1Target_31" AT %Q615.7 : Bool;
   "e1Target_Word" AT %QD612 : DWord;
   "moveCodeKuka" AT %QW616 : Word;   // SIGNAL goTrrigger $IN[ 129]
   "rbDone" AT %I624.0 : Bool;   // SIGNAL rbDoneEdge $OUT[193]
   "x1Target_Word" AT %QD600 : DWord;
   "y1Target_Word" AT %QD604 : DWord;
   "z1Target_Word" AT %QD608 : DWord;
END_VAR
